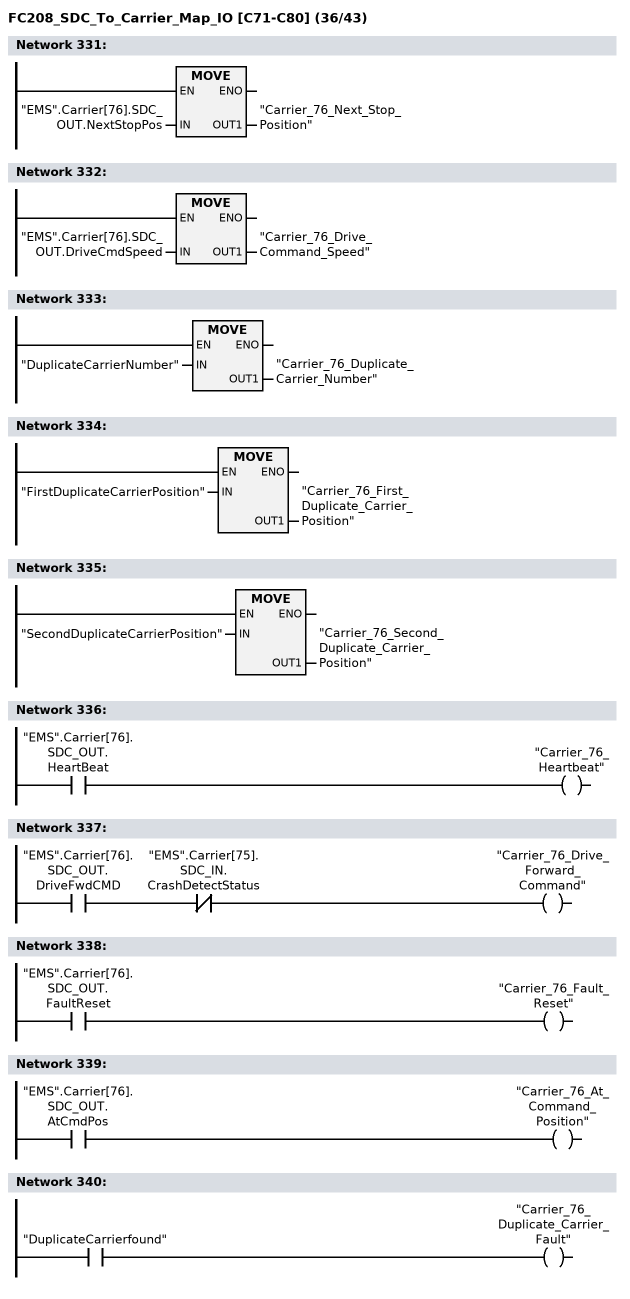
   RUNG wire#powerrail
      Move(in := "EMS".Carrier[76].SDC_OUT.NextStopPos, out1 => "Carrier_76_Next_Stop_Position")
   END_RUNG
   // the same network as SCL:
   "Carrier_76_Next_Stop_Position" := "EMS".Carrier[76].SDC_OUT.NextStopPos;
END_REGION

REGION Network 332
   RUNG wire#powerrail
      Move(in := "EMS".Carrier[76].SDC_OUT.DriveCmdSpeed, out1 => "Carrier_76_Drive_Command_Speed")
   END_RUNG
   // the same network as SCL:
   "Carrier_76_Drive_Command_Speed" := "EMS".Carrier[76].SDC_OUT.DriveCmdSpeed;
END_REGION

REGION Network 333
   RUNG wire#powerrail
      Move(in := "DuplicateCarrierNumber", out1 => "Carrier_76_Duplicate_Carrier_Number")
   END_RUNG
   // the same network as SCL:
   "Carrier_76_Duplicate_Carrier_Number" := "DuplicateCarrierNumber";
END_REGION

REGION Network 334
   RUNG wire#powerrail
      Move(in := "FirstDuplicateCarrierPosition", out1 => "Carrier_76_First_Duplicate_Carrier_Position")
   END_RUNG
   // the same network as SCL:
   "Carrier_76_First_Duplicate_Carrier_Position" := "FirstDuplicateCarrierPosition";
END_REGION

REGION Network 335
   RUNG wire#powerrail
      Move(in := "SecondDuplicateCarrierPosition", out1 => "Carrier_76_Second_Duplicate_Carrier_Position")
   END_RUNG
   // the same network as SCL:
   "Carrier_76_Second_Duplicate_Carrier_Position" := "SecondDuplicateCarrierPosition";
END_REGION

REGION Network 336
   RUNG wire#powerrail
      Contact( "EMS".Carrier[76].SDC_OUT.HeartBeat )
      Coil( "Carrier_76_Heartbeat" )
   END_RUNG
   // the same network as SCL:
   "Carrier_76_Heartbeat" := "EMS".Carrier[76].SDC_OUT.HeartBeat;
END_REGION

REGION Network 337
   RUNG wire#powerrail
      Contact( "EMS".Carrier[76].SDC_OUT.DriveFwdCMD )
      I_Contact( "EMS".Carrier[75].SDC_IN.CrashDetectStatus )
      Coil( "Carrier_76_Drive_Forward_Command" )
   END_RUNG
   // the same network as SCL:
   "Carrier_76_Drive_Forward_Command" := "EMS".Carrier[76].SDC_OUT.DriveFwdCMD AND NOT "EMS".Carrier[75].SDC_IN.CrashDetectStatus;
END_REGION

REGION Network 338
   RUNG wire#powerrail
      Contact( "EMS".Carrier[76].SDC_OUT.FaultReset )
      Coil( "Carrier_76_Fault_Reset" )
   END_RUNG
   // the same network as SCL:
   "Carrier_76_Fault_Reset" := "EMS".Carrier[76].SDC_OUT.FaultReset;
END_REGION

REGION Network 339
   RUNG wire#powerrail
      Contact( "EMS".Carrier[76].SDC_OUT.AtCmdPos )
      Coil( "Carrier_76_At_Command_Position" )
   END_RUNG
   // the same network as SCL:
   "Carrier_76_At_Command_Position" := "EMS".Carrier[76].SDC_OUT.AtCmdPos;
END_REGION

REGION Network 340
   RUNG wire#powerrail
      Contact( "DuplicateCarrierfound" )
      Coil( "Carrier_76_Duplicate_Carrier_Fault" )
   END_RUNG
   // the same network as SCL:
   "Carrier_76_Duplicate_Carrier_Fault" := "DuplicateCarrierfound";
END_REGION

REGION Network 341
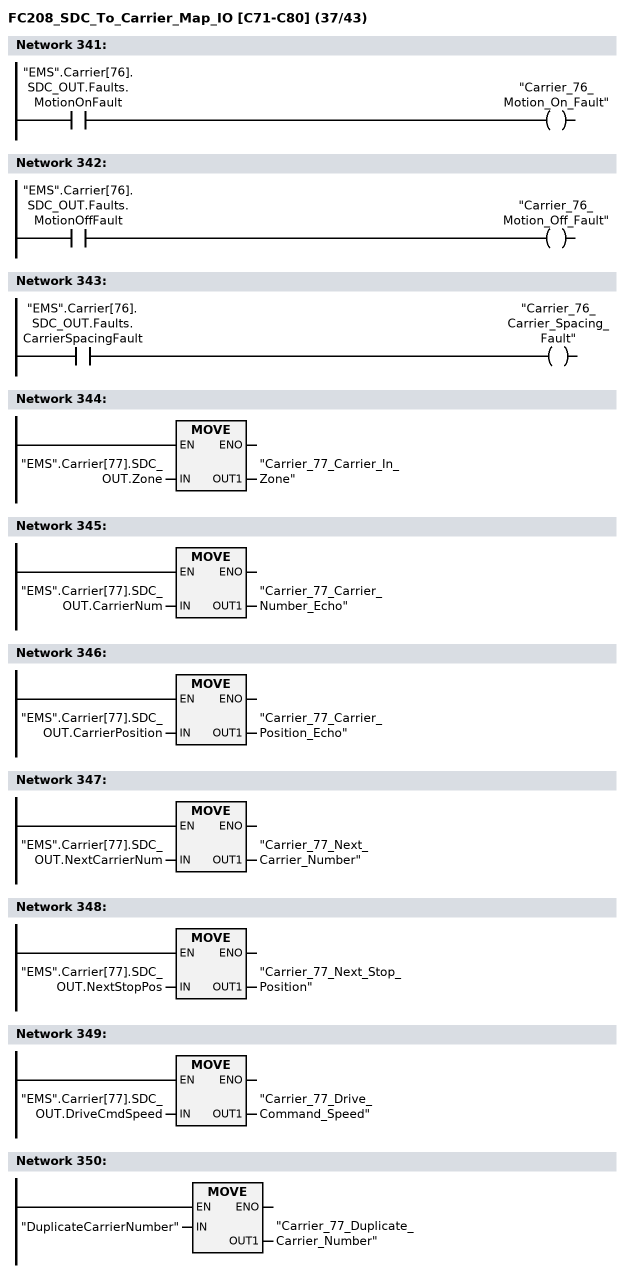
   RUNG wire#powerrail
      Contact( "EMS".Carrier[76].SDC_OUT.Faults.MotionOnFault )
      Coil( "Carrier_76_Motion_On_Fault" )
   END_RUNG
   // the same network as SCL:
   "Carrier_76_Motion_On_Fault" := "EMS".Carrier[76].SDC_OUT.Faults.MotionOnFault;
END_REGION

REGION Network 342
   RUNG wire#powerrail
      Contact( "EMS".Carrier[76].SDC_OUT.Faults.MotionOffFault )
      Coil( "Carrier_76_Motion_Off_Fault" )
   END_RUNG
   // the same network as SCL:
   "Carrier_76_Motion_Off_Fault" := "EMS".Carrier[76].SDC_OUT.Faults.MotionOffFault;
END_REGION

REGION Network 343
   RUNG wire#powerrail
      Contact( "EMS".Carrier[76].SDC_OUT.Faults.CarrierSpacingFault )
      Coil( "Carrier_76_Carrier_Spacing_Fault" )
   END_RUNG
   // the same network as SCL:
   "Carrier_76_Carrier_Spacing_Fault" := "EMS".Carrier[76].SDC_OUT.Faults.CarrierSpacingFault;
END_REGION

REGION Network 344
   RUNG wire#powerrail
      Move(in := "EMS".Carrier[77].SDC_OUT.Zone, out1 => "Carrier_77_Carrier_In_Zone")
   END_RUNG
   // the same network as SCL:
   "Carrier_77_Carrier_In_Zone" := "EMS".Carrier[77].SDC_OUT.Zone;
END_REGION

REGION Network 345
   RUNG wire#powerrail
      Move(in := "EMS".Carrier[77].SDC_OUT.CarrierNum, out1 => "Carrier_77_Carrier_Number_Echo")
   END_RUNG
   // the same network as SCL:
   "Carrier_77_Carrier_Number_Echo" := "EMS".Carrier[77].SDC_OUT.CarrierNum;
END_REGION

REGION Network 346
   RUNG wire#powerrail
      Move(in := "EMS".Carrier[77].SDC_OUT.CarrierPosition, out1 => "Carrier_77_Carrier_Position_Echo")
   END_RUNG
   // the same network as SCL:
   "Carrier_77_Carrier_Position_Echo" := "EMS".Carrier[77].SDC_OUT.CarrierPosition;
END_REGION

REGION Network 347
   RUNG wire#powerrail
      Move(in := "EMS".Carrier[77].SDC_OUT.NextCarrierNum, out1 => "Carrier_77_Next_Carrier_Number")
   END_RUNG
   // the same network as SCL:
   "Carrier_77_Next_Carrier_Number" := "EMS".Carrier[77].SDC_OUT.NextCarrierNum;
END_REGION

REGION Network 348
   RUNG wire#powerrail
      Move(in := "EMS".Carrier[77].SDC_OUT.NextStopPos, out1 => "Carrier_77_Next_Stop_Position")
   END_RUNG
   // the same network as SCL:
   "Carrier_77_Next_Stop_Position" := "EMS".Carrier[77].SDC_OUT.NextStopPos;
END_REGION

REGION Network 349
   RUNG wire#powerrail
      Move(in := "EMS".Carrier[77].SDC_OUT.DriveCmdSpeed, out1 => "Carrier_77_Drive_Command_Speed")
   END_RUNG
   // the same network as SCL:
   "Carrier_77_Drive_Command_Speed" := "EMS".Carrier[77].SDC_OUT.DriveCmdSpeed;
END_REGION

REGION Network 350
   RUNG wire#powerrail
      Move(in := "DuplicateCarrierNumber", out1 => "Carrier_77_Duplicate_Carrier_Number")
   END_RUNG
   // the same network as SCL:
   "Carrier_77_Duplicate_Carrier_Number" := "DuplicateCarrierNumber";
END_REGION

REGION Network 351
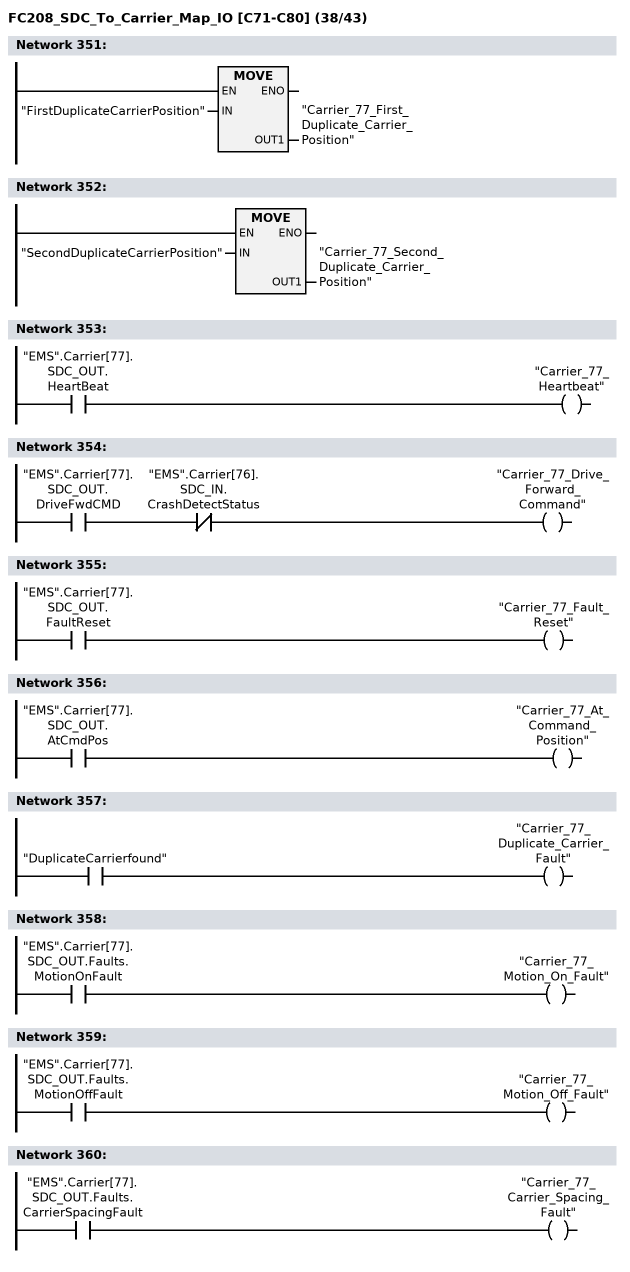
   RUNG wire#powerrail
      Move(in := "FirstDuplicateCarrierPosition", out1 => "Carrier_77_First_Duplicate_Carrier_Position")
   END_RUNG
   // the same network as SCL:
   "Carrier_77_First_Duplicate_Carrier_Position" := "FirstDuplicateCarrierPosition";
END_REGION

REGION Network 352
   RUNG wire#powerrail
      Move(in := "SecondDuplicateCarrierPosition", out1 => "Carrier_77_Second_Duplicate_Carrier_Position")
   END_RUNG
   // the same network as SCL:
   "Carrier_77_Second_Duplicate_Carrier_Position" := "SecondDuplicateCarrierPosition";
END_REGION

REGION Network 353
   RUNG wire#powerrail
      Contact( "EMS".Carrier[77].SDC_OUT.HeartBeat )
      Coil( "Carrier_77_Heartbeat" )
   END_RUNG
   // the same network as SCL:
   "Carrier_77_Heartbeat" := "EMS".Carrier[77].SDC_OUT.HeartBeat;
END_REGION

REGION Network 354
   RUNG wire#powerrail
      Contact( "EMS".Carrier[77].SDC_OUT.DriveFwdCMD )
      I_Contact( "EMS".Carrier[76].SDC_IN.CrashDetectStatus )
      Coil( "Carrier_77_Drive_Forward_Command" )
   END_RUNG
   // the same network as SCL:
   "Carrier_77_Drive_Forward_Command" := "EMS".Carrier[77].SDC_OUT.DriveFwdCMD AND NOT "EMS".Carrier[76].SDC_IN.CrashDetectStatus;
END_REGION

REGION Network 355
   RUNG wire#powerrail
      Contact( "EMS".Carrier[77].SDC_OUT.FaultReset )
      Coil( "Carrier_77_Fault_Reset" )
   END_RUNG
   // the same network as SCL:
   "Carrier_77_Fault_Reset" := "EMS".Carrier[77].SDC_OUT.FaultReset;
END_REGION

REGION Network 356
   RUNG wire#powerrail
      Contact( "EMS".Carrier[77].SDC_OUT.AtCmdPos )
      Coil( "Carrier_77_At_Command_Position" )
   END_RUNG
   // the same network as SCL:
   "Carrier_77_At_Command_Position" := "EMS".Carrier[77].SDC_OUT.AtCmdPos;
END_REGION

REGION Network 357
   RUNG wire#powerrail
      Contact( "DuplicateCarrierfound" )
      Coil( "Carrier_77_Duplicate_Carrier_Fault" )
   END_RUNG
   // the same network as SCL:
   "Carrier_77_Duplicate_Carrier_Fault" := "DuplicateCarrierfound";
END_REGION

REGION Network 358
   RUNG wire#powerrail
      Contact( "EMS".Carrier[77].SDC_OUT.Faults.MotionOnFault )
      Coil( "Carrier_77_Motion_On_Fault" )
   END_RUNG
   // the same network as SCL:
   "Carrier_77_Motion_On_Fault" := "EMS".Carrier[77].SDC_OUT.Faults.MotionOnFault;
END_REGION

REGION Network 359
   RUNG wire#powerrail
      Contact( "EMS".Carrier[77].SDC_OUT.Faults.MotionOffFault )
      Coil( "Carrier_77_Motion_Off_Fault" )
   END_RUNG
   // the same network as SCL:
   "Carrier_77_Motion_Off_Fault" := "EMS".Carrier[77].SDC_OUT.Faults.MotionOffFault;
END_REGION

REGION Network 360
   RUNG wire#powerrail
      Contact( "EMS".Carrier[77].SDC_OUT.Faults.CarrierSpacingFault )
      Coil( "Carrier_77_Carrier_Spacing_Fault" )
   END_RUNG
   // the same network as SCL:
   "Carrier_77_Carrier_Spacing_Fault" := "EMS".Carrier[77].SDC_OUT.Faults.CarrierSpacingFault;
END_REGION

REGION Network 361
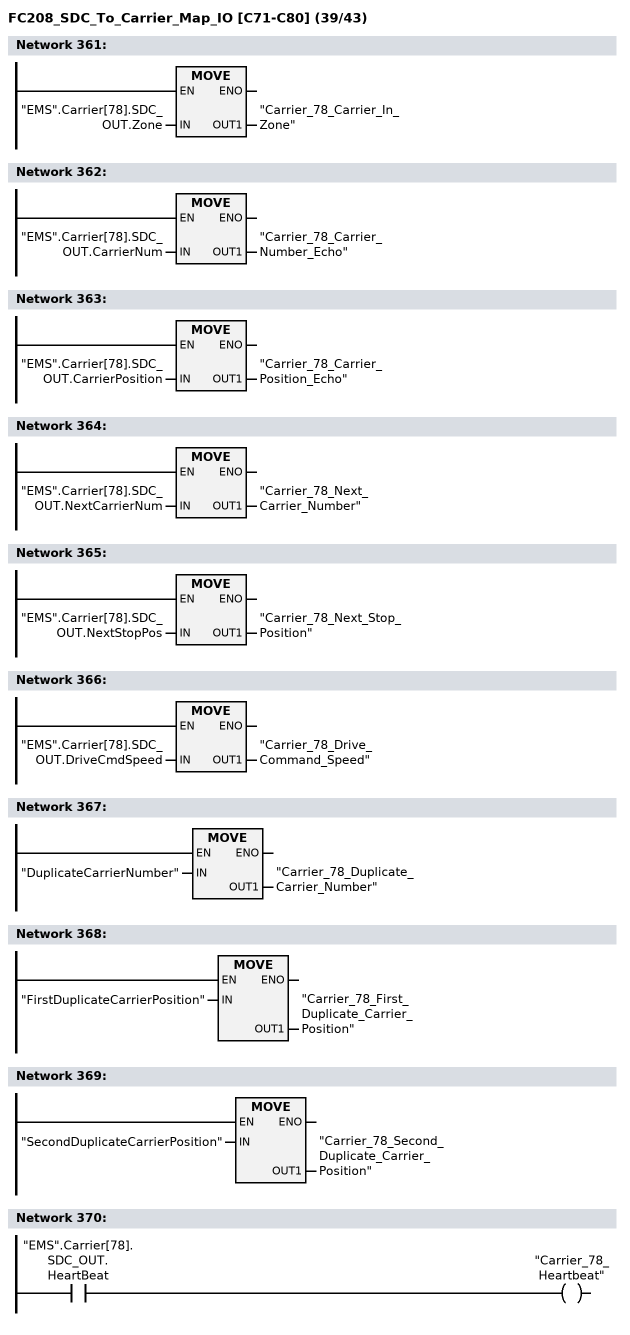
   RUNG wire#powerrail
      Move(in := "EMS".Carrier[78].SDC_OUT.Zone, out1 => "Carrier_78_Carrier_In_Zone")
   END_RUNG
   // the same network as SCL:
   "Carrier_78_Carrier_In_Zone" := "EMS".Carrier[78].SDC_OUT.Zone;
END_REGION

REGION Network 362
   RUNG wire#powerrail
      Move(in := "EMS".Carrier[78].SDC_OUT.CarrierNum, out1 => "Carrier_78_Carrier_Number_Echo")
   END_RUNG
   // the same network as SCL:
   "Carrier_78_Carrier_Number_Echo" := "EMS".Carrier[78].SDC_OUT.CarrierNum;
END_REGION

REGION Network 363
   RUNG wire#powerrail
      Move(in := "EMS".Carrier[78].SDC_OUT.CarrierPosition, out1 => "Carrier_78_Carrier_Position_Echo")
   END_RUNG
   // the same network as SCL:
   "Carrier_78_Carrier_Position_Echo" := "EMS".Carrier[78].SDC_OUT.CarrierPosition;
END_REGION

REGION Network 364
   RUNG wire#powerrail
      Move(in := "EMS".Carrier[78].SDC_OUT.NextCarrierNum, out1 => "Carrier_78_Next_Carrier_Number")
   END_RUNG
   // the same network as SCL:
   "Carrier_78_Next_Carrier_Number" := "EMS".Carrier[78].SDC_OUT.NextCarrierNum;
END_REGION

REGION Network 365
   RUNG wire#powerrail
      Move(in := "EMS".Carrier[78].SDC_OUT.NextStopPos, out1 => "Carrier_78_Next_Stop_Position")
   END_RUNG
   // the same network as SCL:
   "Carrier_78_Next_Stop_Position" := "EMS".Carrier[78].SDC_OUT.NextStopPos;
END_REGION

REGION Network 366
   RUNG wire#powerrail
      Move(in := "EMS".Carrier[78].SDC_OUT.DriveCmdSpeed, out1 => "Carrier_78_Drive_Command_Speed")
   END_RUNG
   // the same network as SCL:
   "Carrier_78_Drive_Command_Speed" := "EMS".Carrier[78].SDC_OUT.DriveCmdSpeed;
END_REGION

REGION Network 367
   RUNG wire#powerrail
      Move(in := "DuplicateCarrierNumber", out1 => "Carrier_78_Duplicate_Carrier_Number")
   END_RUNG
   // the same network as SCL:
   "Carrier_78_Duplicate_Carrier_Number" := "DuplicateCarrierNumber";
END_REGION

REGION Network 368
   RUNG wire#powerrail
      Move(in := "FirstDuplicateCarrierPosition", out1 => "Carrier_78_First_Duplicate_Carrier_Position")
   END_RUNG
   // the same network as SCL:
   "Carrier_78_First_Duplicate_Carrier_Position" := "FirstDuplicateCarrierPosition";
END_REGION

REGION Network 369
   RUNG wire#powerrail
      Move(in := "SecondDuplicateCarrierPosition", out1 => "Carrier_78_Second_Duplicate_Carrier_Position")
   END_RUNG
   // the same network as SCL:
   "Carrier_78_Second_Duplicate_Carrier_Position" := "SecondDuplicateCarrierPosition";
END_REGION

REGION Network 370
   RUNG wire#powerrail
      Contact( "EMS".Carrier[78].SDC_OUT.HeartBeat )
      Coil( "Carrier_78_Heartbeat" )
   END_RUNG
   // the same network as SCL:
   "Carrier_78_Heartbeat" := "EMS".Carrier[78].SDC_OUT.HeartBeat;
END_REGION

REGION Network 371
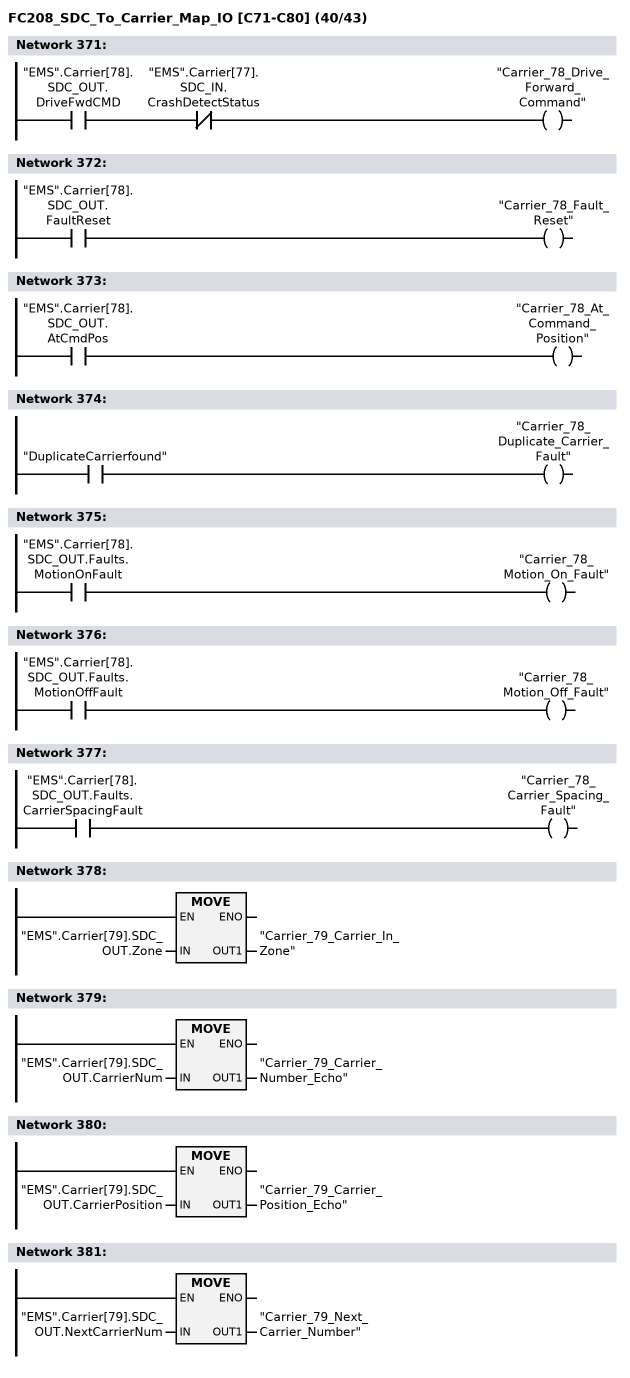
   RUNG wire#powerrail
      Contact( "EMS".Carrier[78].SDC_OUT.DriveFwdCMD )
      I_Contact( "EMS".Carrier[77].SDC_IN.CrashDetectStatus )
      Coil( "Carrier_78_Drive_Forward_Command" )
   END_RUNG
   // the same network as SCL:
   "Carrier_78_Drive_Forward_Command" := "EMS".Carrier[78].SDC_OUT.DriveFwdCMD AND NOT "EMS".Carrier[77].SDC_IN.CrashDetectStatus;
END_REGION

REGION Network 372
   RUNG wire#powerrail
      Contact( "EMS".Carrier[78].SDC_OUT.FaultReset )
      Coil( "Carrier_78_Fault_Reset" )
   END_RUNG
   // the same network as SCL:
   "Carrier_78_Fault_Reset" := "EMS".Carrier[78].SDC_OUT.FaultReset;
END_REGION

REGION Network 373
   RUNG wire#powerrail
      Contact( "EMS".Carrier[78].SDC_OUT.AtCmdPos )
      Coil( "Carrier_78_At_Command_Position" )
   END_RUNG
   // the same network as SCL:
   "Carrier_78_At_Command_Position" := "EMS".Carrier[78].SDC_OUT.AtCmdPos;
END_REGION

REGION Network 374
   RUNG wire#powerrail
      Contact( "DuplicateCarrierfound" )
      Coil( "Carrier_78_Duplicate_Carrier_Fault" )
   END_RUNG
   // the same network as SCL:
   "Carrier_78_Duplicate_Carrier_Fault" := "DuplicateCarrierfound";
END_REGION

REGION Network 375
   RUNG wire#powerrail
      Contact( "EMS".Carrier[78].SDC_OUT.Faults.MotionOnFault )
      Coil( "Carrier_78_Motion_On_Fault" )
   END_RUNG
   // the same network as SCL:
   "Carrier_78_Motion_On_Fault" := "EMS".Carrier[78].SDC_OUT.Faults.MotionOnFault;
END_REGION

REGION Network 376
   RUNG wire#powerrail
      Contact( "EMS".Carrier[78].SDC_OUT.Faults.MotionOffFault )
      Coil( "Carrier_78_Motion_Off_Fault" )
   END_RUNG
   // the same network as SCL:
   "Carrier_78_Motion_Off_Fault" := "EMS".Carrier[78].SDC_OUT.Faults.MotionOffFault;
END_REGION

REGION Network 377
   RUNG wire#powerrail
      Contact( "EMS".Carrier[78].SDC_OUT.Faults.CarrierSpacingFault )
      Coil( "Carrier_78_Carrier_Spacing_Fault" )
   END_RUNG
   // the same network as SCL:
   "Carrier_78_Carrier_Spacing_Fault" := "EMS".Carrier[78].SDC_OUT.Faults.CarrierSpacingFault;
END_REGION

REGION Network 378
   RUNG wire#powerrail
      Move(in := "EMS".Carrier[79].SDC_OUT.Zone, out1 => "Carrier_79_Carrier_In_Zone")
   END_RUNG
   // the same network as SCL:
   "Carrier_79_Carrier_In_Zone" := "EMS".Carrier[79].SDC_OUT.Zone;
END_REGION

REGION Network 379
   RUNG wire#powerrail
      Move(in := "EMS".Carrier[79].SDC_OUT.CarrierNum, out1 => "Carrier_79_Carrier_Number_Echo")
   END_RUNG
   // the same network as SCL:
   "Carrier_79_Carrier_Number_Echo" := "EMS".Carrier[79].SDC_OUT.CarrierNum;
END_REGION

REGION Network 380
   RUNG wire#powerrail
      Move(in := "EMS".Carrier[79].SDC_OUT.CarrierPosition, out1 => "Carrier_79_Carrier_Position_Echo")
   END_RUNG
   // the same network as SCL:
   "Carrier_79_Carrier_Position_Echo" := "EMS".Carrier[79].SDC_OUT.CarrierPosition;
END_REGION

REGION Network 381
   RUNG wire#powerrail
      Move(in := "EMS".Carrier[79].SDC_OUT.NextCarrierNum, out1 => "Carrier_79_Next_Carrier_Number")
   END_RUNG
   // the same network as SCL:
   "Carrier_79_Next_Carrier_Number" := "EMS".Carrier[79].SDC_OUT.NextCarrierNum;
END_REGION

REGION Network 382
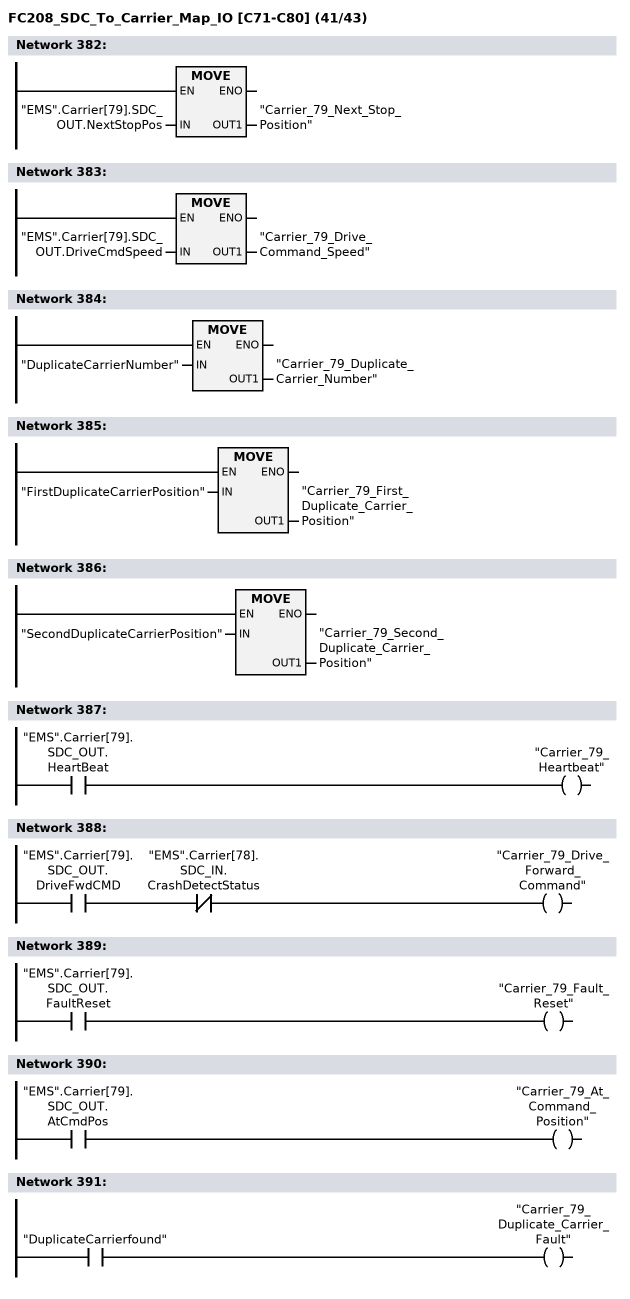
   RUNG wire#powerrail
      Move(in := "EMS".Carrier[79].SDC_OUT.NextStopPos, out1 => "Carrier_79_Next_Stop_Position")
   END_RUNG
   // the same network as SCL:
   "Carrier_79_Next_Stop_Position" := "EMS".Carrier[79].SDC_OUT.NextStopPos;
END_REGION

REGION Network 383
   RUNG wire#powerrail
      Move(in := "EMS".Carrier[79].SDC_OUT.DriveCmdSpeed, out1 => "Carrier_79_Drive_Command_Speed")
   END_RUNG
   // the same network as SCL:
   "Carrier_79_Drive_Command_Speed" := "EMS".Carrier[79].SDC_OUT.DriveCmdSpeed;
END_REGION

REGION Network 384
   RUNG wire#powerrail
      Move(in := "DuplicateCarrierNumber", out1 => "Carrier_79_Duplicate_Carrier_Number")
   END_RUNG
   // the same network as SCL:
   "Carrier_79_Duplicate_Carrier_Number" := "DuplicateCarrierNumber";
END_REGION

REGION Network 385
   RUNG wire#powerrail
      Move(in := "FirstDuplicateCarrierPosition", out1 => "Carrier_79_First_Duplicate_Carrier_Position")
   END_RUNG
   // the same network as SCL:
   "Carrier_79_First_Duplicate_Carrier_Position" := "FirstDuplicateCarrierPosition";
END_REGION

REGION Network 386
   RUNG wire#powerrail
      Move(in := "SecondDuplicateCarrierPosition", out1 => "Carrier_79_Second_Duplicate_Carrier_Position")
   END_RUNG
   // the same network as SCL:
   "Carrier_79_Second_Duplicate_Carrier_Position" := "SecondDuplicateCarrierPosition";
END_REGION

REGION Network 387
   RUNG wire#powerrail
      Contact( "EMS".Carrier[79].SDC_OUT.HeartBeat )
      Coil( "Carrier_79_Heartbeat" )
   END_RUNG
   // the same network as SCL:
   "Carrier_79_Heartbeat" := "EMS".Carrier[79].SDC_OUT.HeartBeat;
END_REGION

REGION Network 388
   RUNG wire#powerrail
      Contact( "EMS".Carrier[79].SDC_OUT.DriveFwdCMD )
      I_Contact( "EMS".Carrier[78].SDC_IN.CrashDetectStatus )
      Coil( "Carrier_79_Drive_Forward_Command" )
   END_RUNG
   // the same network as SCL:
   "Carrier_79_Drive_Forward_Command" := "EMS".Carrier[79].SDC_OUT.DriveFwdCMD AND NOT "EMS".Carrier[78].SDC_IN.CrashDetectStatus;
END_REGION

REGION Network 389
   RUNG wire#powerrail
      Contact( "EMS".Carrier[79].SDC_OUT.FaultReset )
      Coil( "Carrier_79_Fault_Reset" )
   END_RUNG
   // the same network as SCL:
   "Carrier_79_Fault_Reset" := "EMS".Carrier[79].SDC_OUT.FaultReset;
END_REGION

REGION Network 390
   RUNG wire#powerrail
      Contact( "EMS".Carrier[79].SDC_OUT.AtCmdPos )
      Coil( "Carrier_79_At_Command_Position" )
   END_RUNG
   // the same network as SCL:
   "Carrier_79_At_Command_Position" := "EMS".Carrier[79].SDC_OUT.AtCmdPos;
END_REGION

REGION Network 391
   RUNG wire#powerrail
      Contact( "DuplicateCarrierfound" )
      Coil( "Carrier_79_Duplicate_Carrier_Fault" )
   END_RUNG
   // the same network as SCL:
   "Carrier_79_Duplicate_Carrier_Fault" := "DuplicateCarrierfound";
END_REGION

REGION Network 392
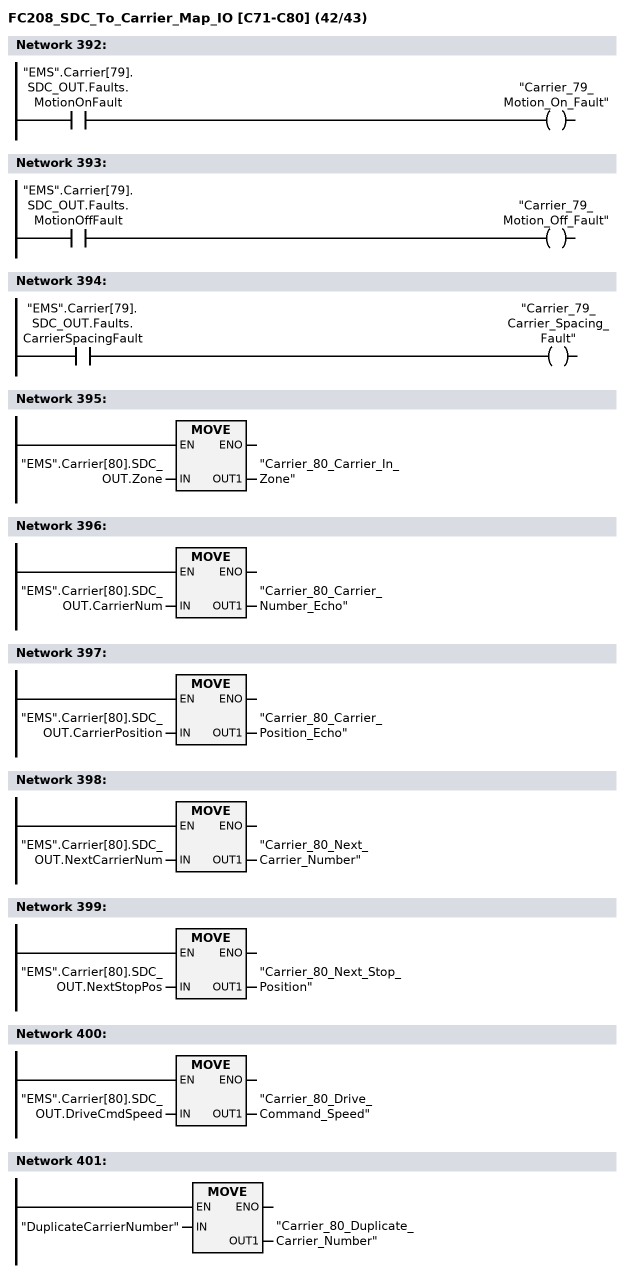
   RUNG wire#powerrail
      Contact( "EMS".Carrier[79].SDC_OUT.Faults.MotionOnFault )
      Coil( "Carrier_79_Motion_On_Fault" )
   END_RUNG
   // the same network as SCL:
   "Carrier_79_Motion_On_Fault" := "EMS".Carrier[79].SDC_OUT.Faults.MotionOnFault;
END_REGION

REGION Network 393
   RUNG wire#powerrail
      Contact( "EMS".Carrier[79].SDC_OUT.Faults.MotionOffFault )
      Coil( "Carrier_79_Motion_Off_Fault" )
   END_RUNG
   // the same network as SCL:
   "Carrier_79_Motion_Off_Fault" := "EMS".Carrier[79].SDC_OUT.Faults.MotionOffFault;
END_REGION

REGION Network 394
   RUNG wire#powerrail
      Contact( "EMS".Carrier[79].SDC_OUT.Faults.CarrierSpacingFault )
      Coil( "Carrier_79_Carrier_Spacing_Fault" )
   END_RUNG
   // the same network as SCL:
   "Carrier_79_Carrier_Spacing_Fault" := "EMS".Carrier[79].SDC_OUT.Faults.CarrierSpacingFault;
END_REGION

REGION Network 395
   RUNG wire#powerrail
      Move(in := "EMS".Carrier[80].SDC_OUT.Zone, out1 => "Carrier_80_Carrier_In_Zone")
   END_RUNG
   // the same network as SCL:
   "Carrier_80_Carrier_In_Zone" := "EMS".Carrier[80].SDC_OUT.Zone;
END_REGION

REGION Network 396
   RUNG wire#powerrail
      Move(in := "EMS".Carrier[80].SDC_OUT.CarrierNum, out1 => "Carrier_80_Carrier_Number_Echo")
   END_RUNG
   // the same network as SCL:
   "Carrier_80_Carrier_Number_Echo" := "EMS".Carrier[80].SDC_OUT.CarrierNum;
END_REGION

REGION Network 397
   RUNG wire#powerrail
      Move(in := "EMS".Carrier[80].SDC_OUT.CarrierPosition, out1 => "Carrier_80_Carrier_Position_Echo")
   END_RUNG
   // the same network as SCL:
   "Carrier_80_Carrier_Position_Echo" := "EMS".Carrier[80].SDC_OUT.CarrierPosition;
END_REGION

REGION Network 398
   RUNG wire#powerrail
      Move(in := "EMS".Carrier[80].SDC_OUT.NextCarrierNum, out1 => "Carrier_80_Next_Carrier_Number")
   END_RUNG
   // the same network as SCL:
   "Carrier_80_Next_Carrier_Number" := "EMS".Carrier[80].SDC_OUT.NextCarrierNum;
END_REGION

REGION Network 399
   RUNG wire#powerrail
      Move(in := "EMS".Carrier[80].SDC_OUT.NextStopPos, out1 => "Carrier_80_Next_Stop_Position")
   END_RUNG
   // the same network as SCL:
   "Carrier_80_Next_Stop_Position" := "EMS".Carrier[80].SDC_OUT.NextStopPos;
END_REGION

REGION Network 400
   RUNG wire#powerrail
      Move(in := "EMS".Carrier[80].SDC_OUT.DriveCmdSpeed, out1 => "Carrier_80_Drive_Command_Speed")
   END_RUNG
   // the same network as SCL:
   "Carrier_80_Drive_Command_Speed" := "EMS".Carrier[80].SDC_OUT.DriveCmdSpeed;
END_REGION

REGION Network 401
   RUNG wire#powerrail
      Move(in := "DuplicateCarrierNumber", out1 => "Carrier_80_Duplicate_Carrier_Number")
   END_RUNG
   // the same network as SCL:
   "Carrier_80_Duplicate_Carrier_Number" := "DuplicateCarrierNumber";
END_REGION

REGION Network 402
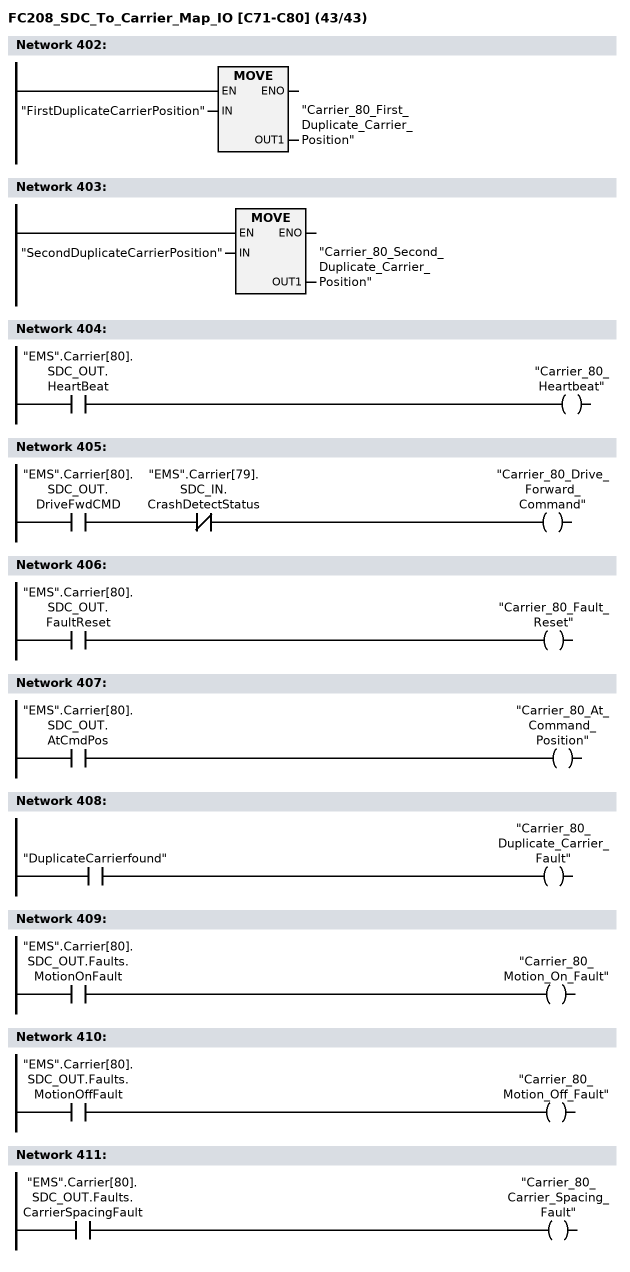
   RUNG wire#powerrail
      Move(in := "FirstDuplicateCarrierPosition", out1 => "Carrier_80_First_Duplicate_Carrier_Position")
   END_RUNG
   // the same network as SCL:
   "Carrier_80_First_Duplicate_Carrier_Position" := "FirstDuplicateCarrierPosition";
END_REGION

REGION Network 403
   RUNG wire#powerrail
      Move(in := "SecondDuplicateCarrierPosition", out1 => "Carrier_80_Second_Duplicate_Carrier_Position")
   END_RUNG
   // the same network as SCL:
   "Carrier_80_Second_Duplicate_Carrier_Position" := "SecondDuplicateCarrierPosition";
END_REGION

REGION Network 404
   RUNG wire#powerrail
      Contact( "EMS".Carrier[80].SDC_OUT.HeartBeat )
      Coil( "Carrier_80_Heartbeat" )
   END_RUNG
   // the same network as SCL:
   "Carrier_80_Heartbeat" := "EMS".Carrier[80].SDC_OUT.HeartBeat;
END_REGION

REGION Network 405
   RUNG wire#powerrail
      Contact( "EMS".Carrier[80].SDC_OUT.DriveFwdCMD )
      I_Contact( "EMS".Carrier[79].SDC_IN.CrashDetectStatus )
      Coil( "Carrier_80_Drive_Forward_Command" )
   END_RUNG
   // the same network as SCL:
   "Carrier_80_Drive_Forward_Command" := "EMS".Carrier[80].SDC_OUT.DriveFwdCMD AND NOT "EMS".Carrier[79].SDC_IN.CrashDetectStatus;
END_REGION

REGION Network 406
   RUNG wire#powerrail
      Contact( "EMS".Carrier[80].SDC_OUT.FaultReset )
      Coil( "Carrier_80_Fault_Reset" )
   END_RUNG
   // the same network as SCL:
   "Carrier_80_Fault_Reset" := "EMS".Carrier[80].SDC_OUT.FaultReset;
END_REGION

REGION Network 407
   RUNG wire#powerrail
      Contact( "EMS".Carrier[80].SDC_OUT.AtCmdPos )
      Coil( "Carrier_80_At_Command_Position" )
   END_RUNG
   // the same network as SCL:
   "Carrier_80_At_Command_Position" := "EMS".Carrier[80].SDC_OUT.AtCmdPos;
END_REGION

REGION Network 408
   RUNG wire#powerrail
      Contact( "DuplicateCarrierfound" )
      Coil( "Carrier_80_Duplicate_Carrier_Fault" )
   END_RUNG
   // the same network as SCL:
   "Carrier_80_Duplicate_Carrier_Fault" := "DuplicateCarrierfound";
END_REGION

REGION Network 409
   RUNG wire#powerrail
      Contact( "EMS".Carrier[80].SDC_OUT.Faults.MotionOnFault )
      Coil( "Carrier_80_Motion_On_Fault" )
   END_RUNG
   // the same network as SCL:
   "Carrier_80_Motion_On_Fault" := "EMS".Carrier[80].SDC_OUT.Faults.MotionOnFault;
END_REGION

REGION Network 410
   RUNG wire#powerrail
      Contact( "EMS".Carrier[80].SDC_OUT.Faults.MotionOffFault )
      Coil( "Carrier_80_Motion_Off_Fault" )
   END_RUNG
   // the same network as SCL:
   "Carrier_80_Motion_Off_Fault" := "EMS".Carrier[80].SDC_OUT.Faults.MotionOffFault;
END_REGION

REGION Network 411
   RUNG wire#powerrail
      Contact( "EMS".Carrier[80].SDC_OUT.Faults.CarrierSpacingFault )
      Coil( "Carrier_80_Carrier_Spacing_Fault" )
   END_RUNG
   // the same network as SCL:
   "Carrier_80_Carrier_Spacing_Fault" := "EMS".Carrier[80].SDC_OUT.Faults.CarrierSpacingFault;
END_REGION
END_FUNCTION

FUNCTION "FC209_SDC_To_Carrier_Map_IO [C81-C82]" : Void   // FC209, LAD
{ S7_Optimized_Access := 'TRUE' }
VERSION : 0.1
BEGIN

REGION Network 1
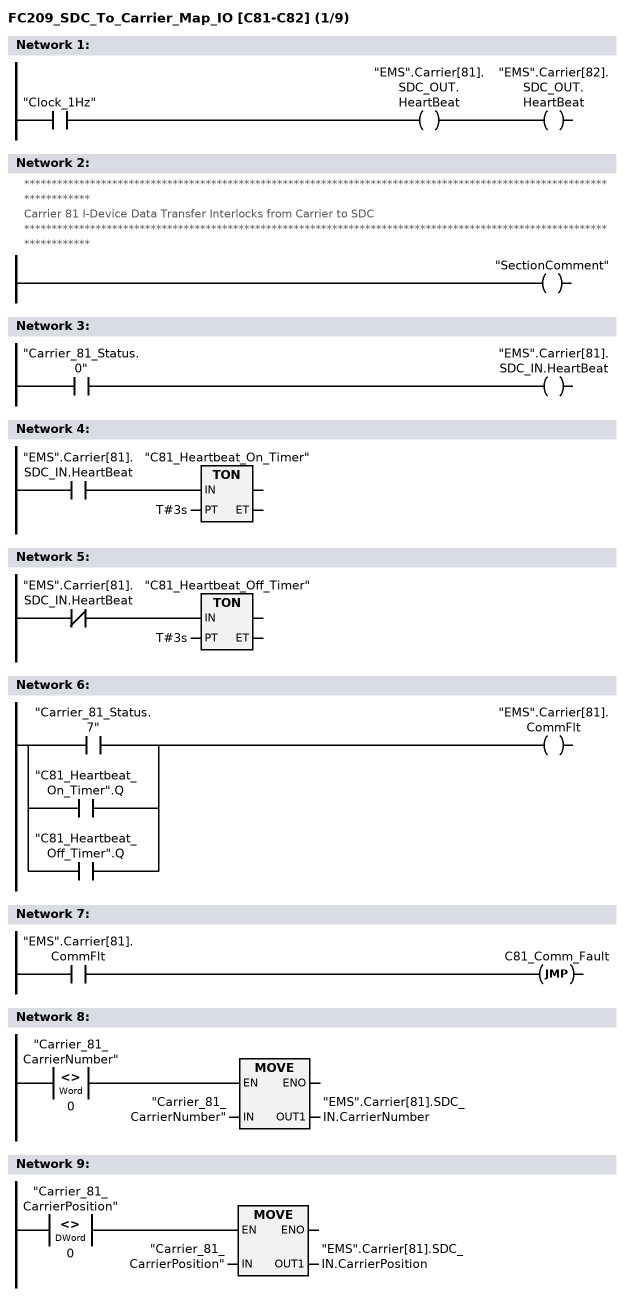
   RUNG wire#powerrail
      Contact( "Clock_1Hz" )
      Coil( "EMS".Carrier[81].SDC_OUT.HeartBeat )
      Coil( "EMS".Carrier[82].SDC_OUT.HeartBeat )
   END_RUNG
   // the same network as SCL:
   "EMS".Carrier[81].SDC_OUT.HeartBeat := "Clock_1Hz";
   "EMS".Carrier[82].SDC_OUT.HeartBeat := "Clock_1Hz";
END_REGION
